// TIA Portal project "HydroPlantProject_V15.1" (V15.1) (continued)

   //EStop Alarm
   IF NOT "EStop" AND NOT "EStopAlarm" THEN
       "EStopAlarm" := 1;
       "EStopNotify" := 1;
   END_IF;

   IF "EStopAlarm" AND "AlarmReset" THEN
       "EStopAlarm" := 0;
       "EStopNotify" := 0;
   END_IF;

   IF "EStopNotify" AND "AlarmSilence" THEN
       "EStopNotify" := 0;
   END_IF;



   //Alarm Horn Control
   IF "FaultMode" AND NOT "AlarmHorn_Ctrl" THEN
       "AlarmHorn_Ctrl" := 1;
   END_IF;

   IF "AlarmHorn_Ctrl" AND ("AlarmReset" OR "AlarmSilence") THEN
       "AlarmHorn_Ctrl" := 0;
   END_IF;
END_FUNCTION_BLOCK

FUNCTION_BLOCK "ALARMS_STL"   // FB13, STL
{ S7_Optimized_Access := 'TRUE' }
VERSION : 0.1
   VAR
      OS1 : Bool;
      OS2 : Bool;
      OS3 : Bool;
      OS4 : Bool;
      OS5 : Bool;
      OS6 : Bool;
      OS7 : Bool;
      OS8 : Bool;
      OS9 : Bool;
      OS10 : Bool;
      OS11 : Bool;
      OS12 : Bool;
      OS13 : Bool;
      OS14 : Bool;
      OS15 : Bool;
      OS16 : Bool;
      OS17 : Bool;
   END_VAR
   VAR_TEMP
      ti1 : Time;
      ti2 : Time;
      ti3 : Time;
      ti4 : Time;
      ti5 : Time;
      ti6 : Time;
      ti7 : Time;
      t1 : Time;
      t2 : Time;
      t3 : Time;
      t4 : Time;
      t5 : Time;
      t6 : Time;
      t7 : Time;
      OILAT : Bool;
      OLFAT : Bool;
      OCAT : Bool;
      HOTAT : Bool;
      OSAT : Bool;
      HOFAT : Bool;
      BFAT : Bool;
   END_VAR
BEGIN

REGION Network 1
   //Oil Low Flow Alarm
         L     "OilFlow";
         L     "OilLLflowSp";
         <I;
         A     "OilPumpVFDen_Out";
         AN    "Brake_Out";
         JC    OLFtimer;
         CLR;
         A     "AlarmReset";
         FP    #OS1;
         JC    ResetOLFalarm;
         CLR;
         A     "AlarmSilence";
         FP    #OS2;
         JC    ResetOLFnotify;
         JU    OvercurrentAlarm;

   OLFtimer:CALL  "CONVERTTIME"
         ( Int1  := "OilLowFlowDelay_Sp",
           Time1 := #ti1
         );
         CALL  TON, "IEC_Timer_0_DB_18"
         ( IN := TRUE,
           PT := #ti1,
           Q  := #OLFAT,
           ET := #t1
         );
         A     #OLFAT;
         JC    SetOLFalarm;
         JU    OvercurrentAlarm;

   SetOLFalarm:SET;
         S     "OilLowFlowAlarm";
         S     "OilLowFlowNotify";
         JU    OvercurrentAlarm;

   ResetOLFalarm:R     "OilLowFlowAlarm";
         R     "OilLowFlowNotify";
         JU    OvercurrentAlarm;

   ResetOLFnotify:R     "OilLowFlowNotify";
         JU    OvercurrentAlarm;


   //Overcurrent Alarm
   OvercurrentAlarm:L     "Current";
         L     "OvercurrentSp";
         >I;
         JC    OCtimer;
         CLR;
         A     "AlarmReset";
         FP    #OS3;
         JC    ResetOCalarm;
         CLR;
         A     "AlarmSilence";
         FP    #OS4;
         JC    ResetOCnotify;
         JU    HighOilTempAlarm;

   OCtimer:CALL  "CONVERTTIME"
         ( Int1  := "OvercurrentDelay_Sp",
           Time1 := #ti2
         );
         CALL  TON, "IEC_Timer_0_DB_19"
         ( IN := true,
           PT := #ti2,
           Q  := #OCAT,
           ET := #t2
         );
         A     #OCAT;
         JC    SetOCalarm;
         JU    HighOilTempAlarm;

   SetOCalarm:SET;
         S     "OvercurrentAlarm";
         S     "OvercurrentNotify";
         JU    HighOilTempAlarm;

   ResetOCalarm:R     "OvercurrentAlarm";
         R     "OvercurrentNotify";
         JU    HighOilTempAlarm;

   ResetOCnotify:R     "OvercurrentNotify";
         JU    HighOilTempAlarm;


   //High Oil Temp Alarm
   HighOilTempAlarm:L     "OilTemp";
         L     "HighOilTempSp";
         >I;
         JC    HOTtimer;
         CLR;
         A     "AlarmReset";
         FP    #OS5;
         JC    ResetHOTalarm;
         CLR;
         A     "AlarmSilence";
         FP    #OS6;
         JC    ResetHOTnotify;
         JU    OverspeedAlarm;

   HOTtimer:CALL  "CONVERTTIME"
         ( Int1  := "HighOilTempDelay_Sp",
           Time1 := #ti3
         );
         CALL  TON, "IEC_Timer_0_DB_20"
         ( IN := TRUE,
           PT := #ti3,
           Q  := #HOTAT,
           ET := #t3
         );
         A     #HOTAT;
         JC    SetHOTalarm;
         JU    OverspeedAlarm;

   SetHOTalarm:SET;
         S     "HighOilTempAlarm";
         S     "HighOilTempNotify";
         JU    OverspeedAlarm;

   ResetHOTalarm:R     "HighOilTempAlarm";
         R     "HighOilTempNotify";
         JU    OverspeedAlarm;

   ResetHOTnotify:R     "HighOilTempNotify";
         JU    OverspeedAlarm;


   //Overspeed Alarm
   OverspeedAlarm:L     "RPM";
         L     "OverspeedSp";
         >I;
         JC    OStimer;
         CLR;
         A     "AlarmReset";
         FP    #OS7;
         JC    ResetOSalarm;
         CLR;
         A     "AlarmSilence";
         FP    #OS8;
         JC    ResetOSnotify;
         JU    HighOilFlowAlarm;

   OStimer:CALL  "CONVERTTIME"
         ( Int1  := "OverspeedDelay_Sp",
           Time1 := #ti4
         );
         CALL  TON, "IEC_Timer_0_DB_21"
         ( IN := TRUE,
           PT := #ti4,
           Q  := #OSAT,
           ET := #t4
         );
         A     #OSAT;
         JC    SetOSalarm;
         JU    HighOilFlowAlarm;

   SetOSalarm:SET;
         S     "OverspeedAlarm";
         S     "OverspeedNotify";
         JU    HighOilFlowAlarm;

   ResetOSalarm:R     "OverspeedAlarm";
         R     "OverspeedNotify";
         JU    HighOilFlowAlarm;

   ResetOSnotify:R     "OverspeedNotify";
         JU    HighOilFlowAlarm;


   //High Oil Flow Alarm
   HighOilFlowAlarm:L     "OilFlow";
         L     "OilHHflowSp";
         >I;
         JC    HOFtimer;
         CLR;
         A     "AlarmReset";
         FP    #OS9;
         JC    ResetHOFalarm;
         CLR;
         A     "AlarmSilence";
         FP    #OS10;
         JC    ResetHOFnotify;
         JU    BrakeFailureAlarm;

   HOFtimer:CALL  "CONVERTTIME"
         ( Int1  := "OilHighFlowDelay_Sp",
           Time1 := #ti5
         );
         CALL  TON, "IEC_Timer_0_DB_22"
         ( IN := TRUE,
           PT := #ti5,
           Q  := #HOFAT,
           ET := #t5
         );
         A     #HOFAT;
         JC    SetHOFalarm;
         JU    BrakeFailureAlarm;

   SetHOFalarm:SET;
         S     "OilHighFlowAlarm";
         S     "OilHighFlowNotify";
         JU    BrakeFailureAlarm;

   ResetHOFalarm:R     "OilHighFlowAlarm";
         R     "OilHighFlowNotify";
         JU    BrakeFailureAlarm;

   ResetHOFnotify:R     "OilHighFlowNotify";
         JU    BrakeFailureAlarm;


   //Brake Failure Alarm
   BrakeFailureAlarm:L     "RPM";
         L     0;
         >I;
         A     "Brake_Out";
         JC    BFtimer;
         CLR;
         A     "AlarmReset";
         FP    #OS11;
         JC    ResetBFalarm;
         CLR;
         A     "AlarmSilence";
         FP    #OS12;
         JC    ResetBFnotify;
         JU    EStoplarm;

   BFtimer:CALL  "CONVERTTIME"
         ( Int1  := "BrakeFailureDelay_Sp",
           Time1 := #ti6
         );
         CALL  TON, "IEC_Timer_0_DB_23"
         ( IN := TRUE,
           PT := #ti6,
           Q  := #BFAT,
           ET :=
         );
         A     #BFAT;
         JC    SetBFalarm;
         JU    EStoplarm;

   SetBFalarm:SET;
         S     "BrakeFailureAlarm";
         S     "BrakeFailureNotify";
         JU    EStoplarm;

   ResetBFalarm:R     "BrakeFailureAlarm";
         R     "BrakeFailureNotify";
         JU    EStoplarm;

   ResetBFnotify:R     "BrakeFailureNotify";
         JU    EStoplarm;


   //EStop Alarm
   EStoplarm:AN    "EStop";
         FP    #OS13;
         JC    SetESalarm;
         CLR;
         A     "AlarmReset";
         FP    #OS14;
         JC    ResetESalarm;
         CLR;
         A     "AlarmSilence";
         FP    #OS15;
         JC    ResetESnotify;
         JU    AlarmHornCtrl;

   SetESalarm:SET;
         S     "EStopAlarm";
         S     "EStopNotify";
         JU    AlarmHornCtrl;

   ResetESalarm:R     "EStopAlarm";
         R     "EStopNotify";
         JU    AlarmHornCtrl;

   ResetESnotify:R     "EStopNotify";
         JU    AlarmHornCtrl;



   //Alarm Horn Control
   AlarmHornCtrl:A     "FaultMode";
         FP    #OS16;
         JC    SetAlarmHorn;
         CLR;
         A     "AlarmReset";
         O     "AlarmSilence";
         FP    #OS17;
         JC    ResetAlarmHorn;
         JU    EndOfLine;

   SetAlarmHorn:SET;
         S     "AlarmHorn_Ctrl";
         JU    EndOfLine;

   ResetAlarmHorn:R     "AlarmHorn_Ctrl";
         JU    EndOfLine;



   EndOfLine:BE;
END_REGION
END_FUNCTION_BLOCK

FUNCTION_BLOCK "MODES_LAD"   // FB14, LAD
{ S7_Optimized_Access := 'TRUE' }
VERSION : 0.1
   VAR
      OS1 : Bool;
      OS2 : Bool;
      OS3 : Bool;
      OS4 : Bool;
      OS5 : Bool;
   END_VAR
   VAR_TEMP
      tv1 : Int;
      ti1 : Time;
      tv2 : Int;
      tv3 : Int;
      tv4 : Int;
      ti2 : Time;
      tv5 : Int;
      ti3 : Time;
   END_VAR
   VAR_TEMP   // added for the SCL form of the ladder/FBD networks
      _w1 : Bool;
      _w2 : Bool;
      _w3 : Bool;
   END_VAR
BEGIN

REGION Network 1
   // Warmup Mode
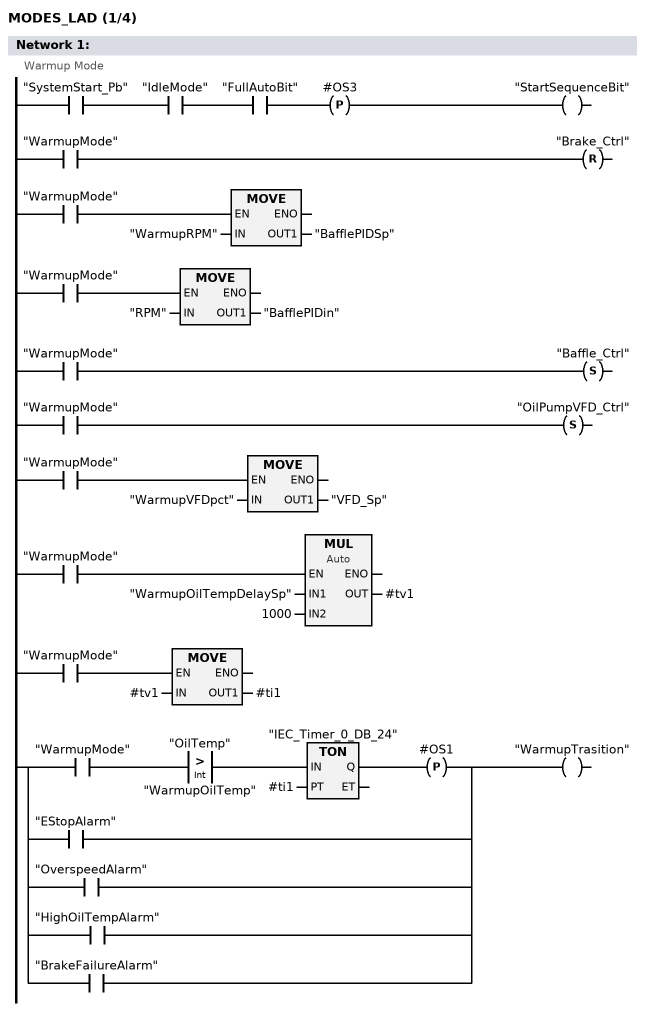
   #_w1 := "SystemStart_Pb" AND "IdleMode" AND "FullAutoBit";
   #_w2 := #_w1 AND NOT #OS3;   // rising edge
   #OS3 := #_w1;
   "StartSequenceBit" := #_w2;
   IF "WarmupMode" THEN
       "Brake_Ctrl" := FALSE;
       "BafflePIDSp" := "WarmupRPM";
       "BafflePIDin" := "RPM";
       "Baffle_Ctrl" := TRUE;
       "OilPumpVFD_Ctrl" := TRUE;
       "VFD_Sp" := "WarmupVFDpct";
       #tv1 := "WarmupOilTempDelaySp" * 1000;
       #ti1 := #tv1;
   END_IF;
   "IEC_Timer_0_DB_24".TON(IN := "WarmupMode" AND ("OilTemp" > "WarmupOilTemp"), PT := #ti1);
   #_w3 := "IEC_Timer_0_DB_24".Q AND NOT #OS1;   // rising edge
   #OS1 := "IEC_Timer_0_DB_24".Q;
   "WarmupTrasition" := #_w3 OR "EStopAlarm" OR "OverspeedAlarm" OR "HighOilTempAlarm" OR "BrakeFailureAlarm";
END_REGION

REGION Network 2
   // Stabilize Mode
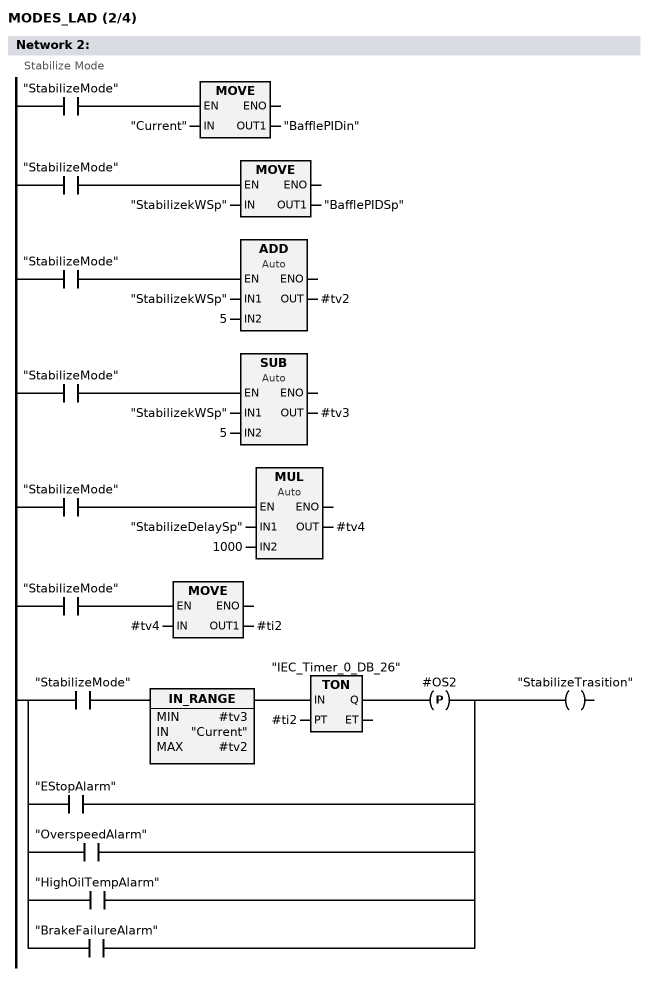
   IF "StabilizeMode" THEN
       "BafflePIDin" := "Current";
       "BafflePIDSp" := "StabilizekWSp";
       #tv2 := "StabilizekWSp" + 5;
       #tv3 := "StabilizekWSp" - 5;
       #tv4 := "StabilizeDelaySp" * 1000;
       #ti2 := #tv4;
   END_IF;
   "IEC_Timer_0_DB_26".TON(IN := "StabilizeMode" AND (#tv3 <= "Current") AND ("Current" <= #tv2), PT := #ti2);
   #_w1 := "IEC_Timer_0_DB_26".Q AND NOT #OS2;   // rising edge
   #OS2 := "IEC_Timer_0_DB_26".Q;
   "StabilizeTrasition" := #_w1 OR "EStopAlarm" OR "OverspeedAlarm" OR "HighOilTempAlarm" OR "BrakeFailureAlarm";
END_REGION

REGION Network 3
   // Generation Mode
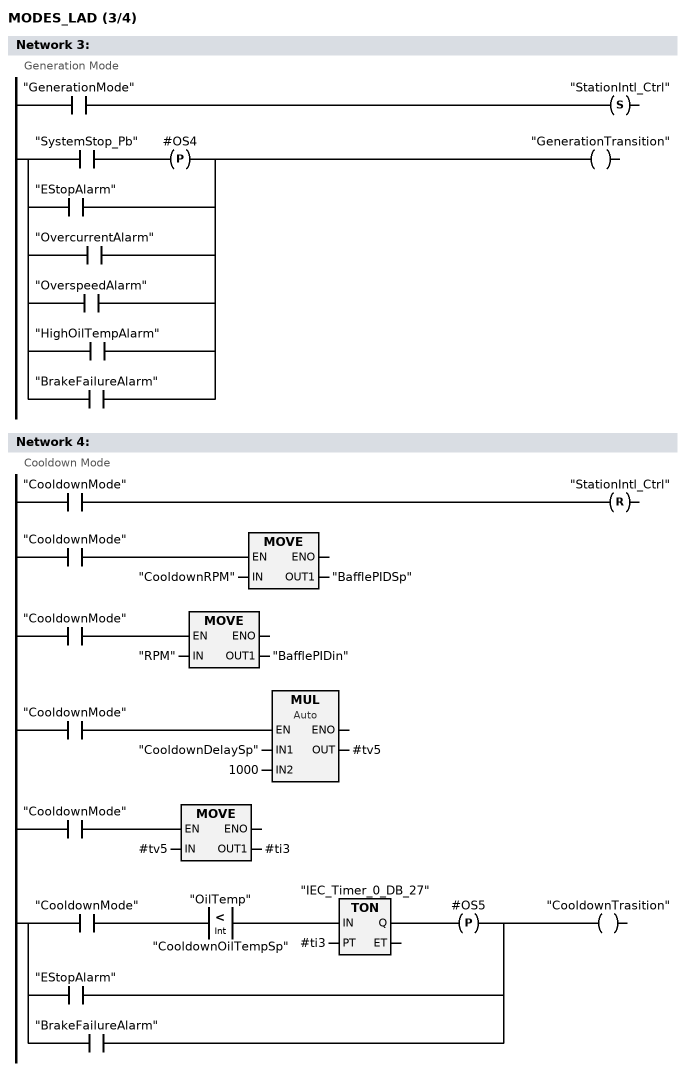
   RUNG wire#powerrail
      Contact( "GenerationMode" )
      S_Coil( "StationIntl_Ctrl" )
   END_RUNG
   RUNG wire#powerrail
      Contact( "SystemStop_Pb" )
      P_Trig( #OS4 )
      wire#w1
      Coil( "GenerationTransition" )
   END_RUNG
   RUNG wire#powerrail
      Contact( "EStopAlarm" )
   END_RUNG wire#w1
   RUNG wire#powerrail
      Contact( "OvercurrentAlarm" )
   END_RUNG wire#w1
   RUNG wire#powerrail
      Contact( "OverspeedAlarm" )
   END_RUNG wire#w1
   RUNG wire#powerrail
      Contact( "HighOilTempAlarm" )
   END_RUNG wire#w1
   RUNG wire#powerrail
      Contact( "BrakeFailureAlarm" )
   END_RUNG wire#w1
   // the same network as SCL:
   IF "GenerationMode" THEN "StationIntl_Ctrl" := TRUE; END_IF;
   #_w1 := "SystemStop_Pb" AND NOT #OS4;   // rising edge
   #OS4 := "SystemStop_Pb";
   "GenerationTransition" := #_w1 OR "EStopAlarm" OR "OvercurrentAlarm" OR "OverspeedAlarm" OR "HighOilTempAlarm" OR "BrakeFailureAlarm";
END_REGION

REGION Network 4
   // Cooldown Mode
   IF "CooldownMode" THEN
       "StationIntl_Ctrl" := FALSE;
       "BafflePIDSp" := "CooldownRPM";
       "BafflePIDin" := "RPM";
       #tv5 := "CooldownDelaySp" * 1000;
       #ti3 := #tv5;
   END_IF;
   "IEC_Timer_0_DB_27".TON(IN := "CooldownMode" AND ("OilTemp" < "CooldownOilTempSp"), PT := #ti3);
   #_w1 := "IEC_Timer_0_DB_27".Q AND NOT #OS5;   // rising edge
   #OS5 := "IEC_Timer_0_DB_27".Q;
   "CooldownTrasition" := #_w1 OR "EStopAlarm" OR "BrakeFailureAlarm";
END_REGION

REGION Network 5
   // Idle Mode
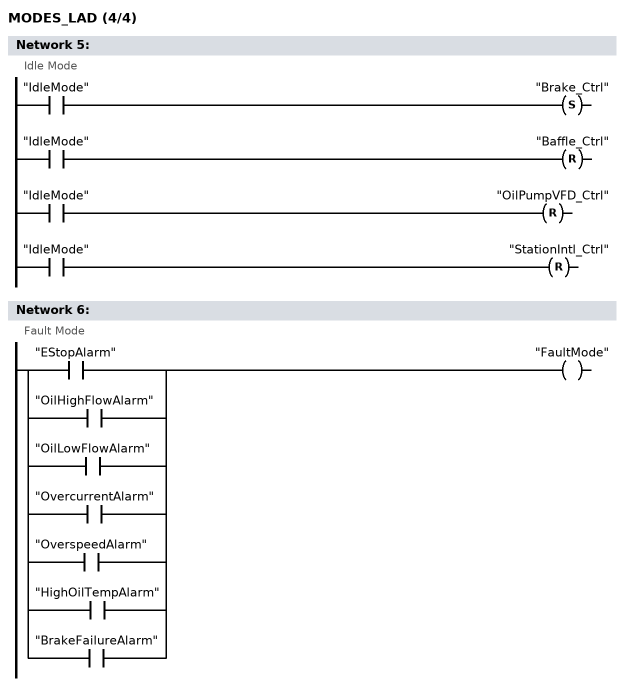
   RUNG wire#powerrail
      Contact( "IdleMode" )
      S_Coil( "Brake_Ctrl" )
   END_RUNG
   RUNG wire#powerrail
      Contact( "IdleMode" )
      R_Coil( "Baffle_Ctrl" )
   END_RUNG
   RUNG wire#powerrail
      Contact( "IdleMode" )
      R_Coil( "OilPumpVFD_Ctrl" )
   END_RUNG
   RUNG wire#powerrail
      Contact( "IdleMode" )
      R_Coil( "StationIntl_Ctrl" )
   END_RUNG
   // the same network as SCL:
   IF "IdleMode" THEN
       "Brake_Ctrl" := TRUE;
       "Baffle_Ctrl" := FALSE;
       "OilPumpVFD_Ctrl" := FALSE;
       "StationIntl_Ctrl" := FALSE;
   END_IF;
END_REGION

REGION Network 6
   // Fault Mode
   RUNG wire#powerrail
      Contact( "EStopAlarm" )
      wire#w1
      Coil( "FaultMode" )
   END_RUNG
   RUNG wire#powerrail
      Contact( "OilHighFlowAlarm" )
   END_RUNG wire#w1
   RUNG wire#powerrail
      Contact( "OilLowFlowAlarm" )
   END_RUNG wire#w1
   RUNG wire#powerrail
      Contact( "OvercurrentAlarm" )
   END_RUNG wire#w1
   RUNG wire#powerrail
      Contact( "OverspeedAlarm" )
   END_RUNG wire#w1
   RUNG wire#powerrail
      Contact( "HighOilTempAlarm" )
   END_RUNG wire#w1
   RUNG wire#powerrail
      Contact( "BrakeFailureAlarm" )
   END_RUNG wire#w1
   // the same network as SCL:
   "FaultMode" := "EStopAlarm" OR "OilHighFlowAlarm" OR "OilLowFlowAlarm" OR "OvercurrentAlarm" OR "OverspeedAlarm" OR "HighOilTempAlarm" OR "BrakeFailureAlarm";
END_REGION
END_FUNCTION_BLOCK

FUNCTION_BLOCK "MODES_FBD"   // FB15, FBD
{ S7_Optimized_Access := 'TRUE' }
VERSION : 0.1
   VAR
      OS1 : Bool;
      OS2 : Bool;
      OS3 : Bool;
      OS4 : Bool;
      OS5 : Bool;
   END_VAR
   VAR_TEMP
      ti1 : Time;
      tv1 : Int;
      tv2 : Int;
      ti3 : Time;
      ti2 : Time;
   END_VAR
   VAR_TEMP   // added for the SCL form of the ladder/FBD networks
      _w1 : Bool;
      _w2 : Bool;
      _w3 : Bool;
   END_VAR
BEGIN

REGION Network 1
   // Warmup Mode
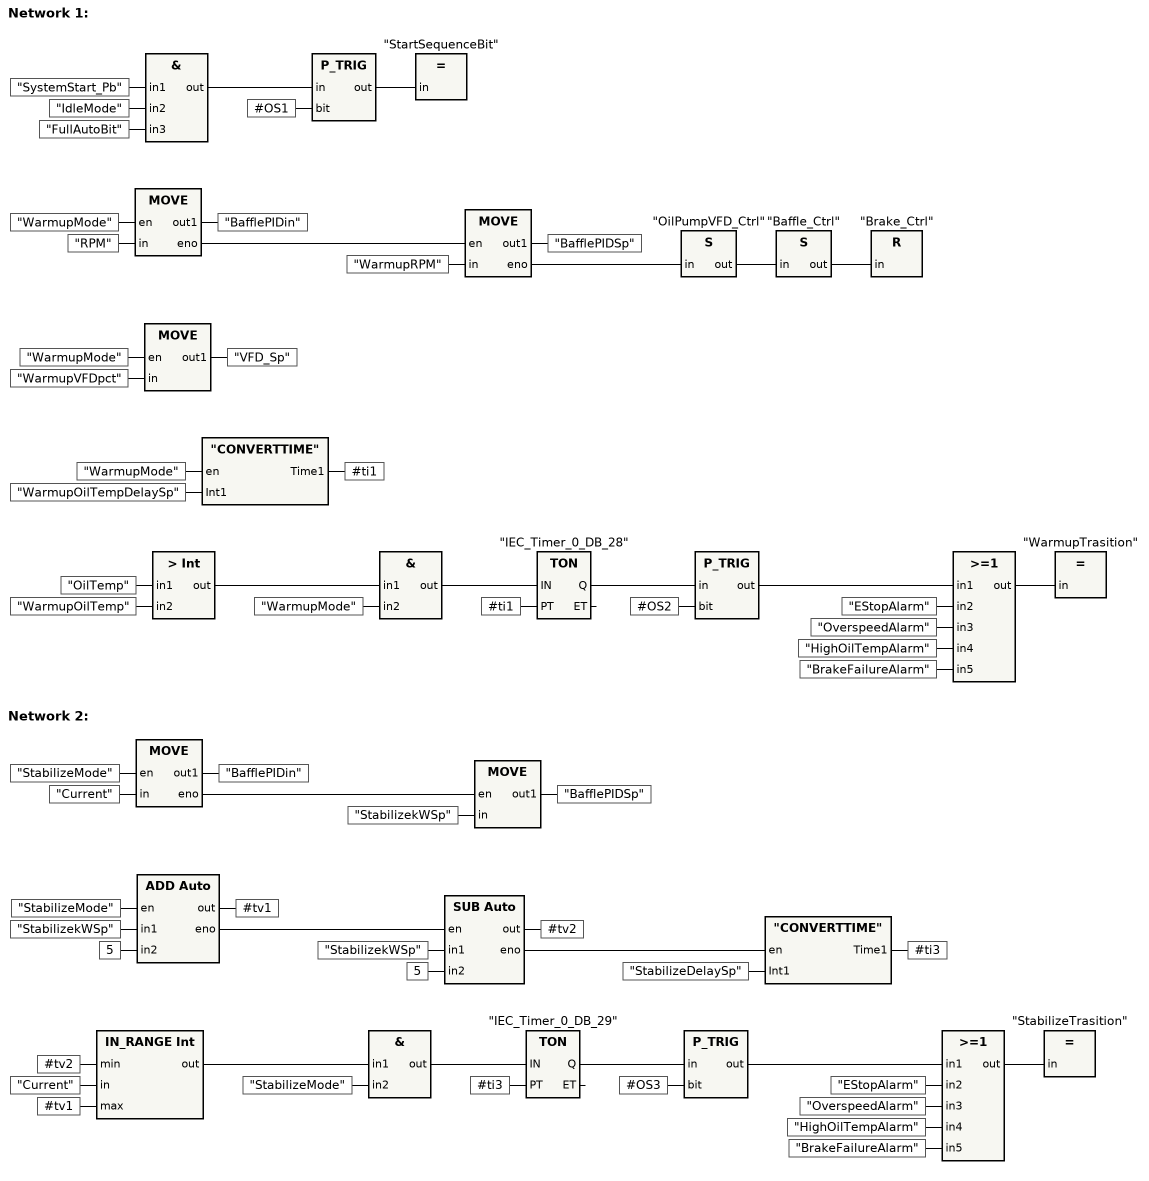
   #_w1 := "SystemStart_Pb" AND "IdleMode" AND "FullAutoBit";
   #_w2 := #_w1 AND NOT #OS1;   // rising edge
   #OS1 := #_w1;
   "StartSequenceBit" := #_w2;
   IF "WarmupMode" THEN
       "BafflePIDin" := "RPM";
       "BafflePIDSp" := "WarmupRPM";
       "OilPumpVFD_Ctrl" := TRUE;
       "Baffle_Ctrl" := TRUE;
       "Brake_Ctrl" := FALSE;
       "VFD_Sp" := "WarmupVFDpct";
       "CONVERTTIME"(Int1 := "WarmupOilTempDelaySp", Time1 => #ti1);
   END_IF;
   "IEC_Timer_0_DB_28".TON(IN := ("OilTemp" > "WarmupOilTemp") AND "WarmupMode", PT := #ti1);
   #_w3 := "IEC_Timer_0_DB_28".Q AND NOT #OS2;   // rising edge
   #OS2 := "IEC_Timer_0_DB_28".Q;
   "WarmupTrasition" := #_w3 OR "EStopAlarm" OR "OverspeedAlarm" OR "HighOilTempAlarm" OR "BrakeFailureAlarm";
END_REGION

REGION Network 2
   // Stabilize Mode
   IF "StabilizeMode" THEN
       "BafflePIDin" := "Current";
       "BafflePIDSp" := "StabilizekWSp";
       #tv1 := "StabilizekWSp" + 5;
       #tv2 := "StabilizekWSp" - 5;
       "CONVERTTIME"(Int1 := "StabilizeDelaySp", Time1 => #ti3);
   END_IF;
   "IEC_Timer_0_DB_29".TON(IN := (#tv2 <= "Current") AND ("Current" <= #tv1) AND "StabilizeMode", PT := #ti3);
   #_w1 := "IEC_Timer_0_DB_29".Q AND NOT #OS3;   // rising edge
   #OS3 := "IEC_Timer_0_DB_29".Q;
   "StabilizeTrasition" := #_w1 OR "EStopAlarm" OR "OverspeedAlarm" OR "HighOilTempAlarm" OR "BrakeFailureAlarm";
END_REGION

REGION Network 3
   // Generation Mode
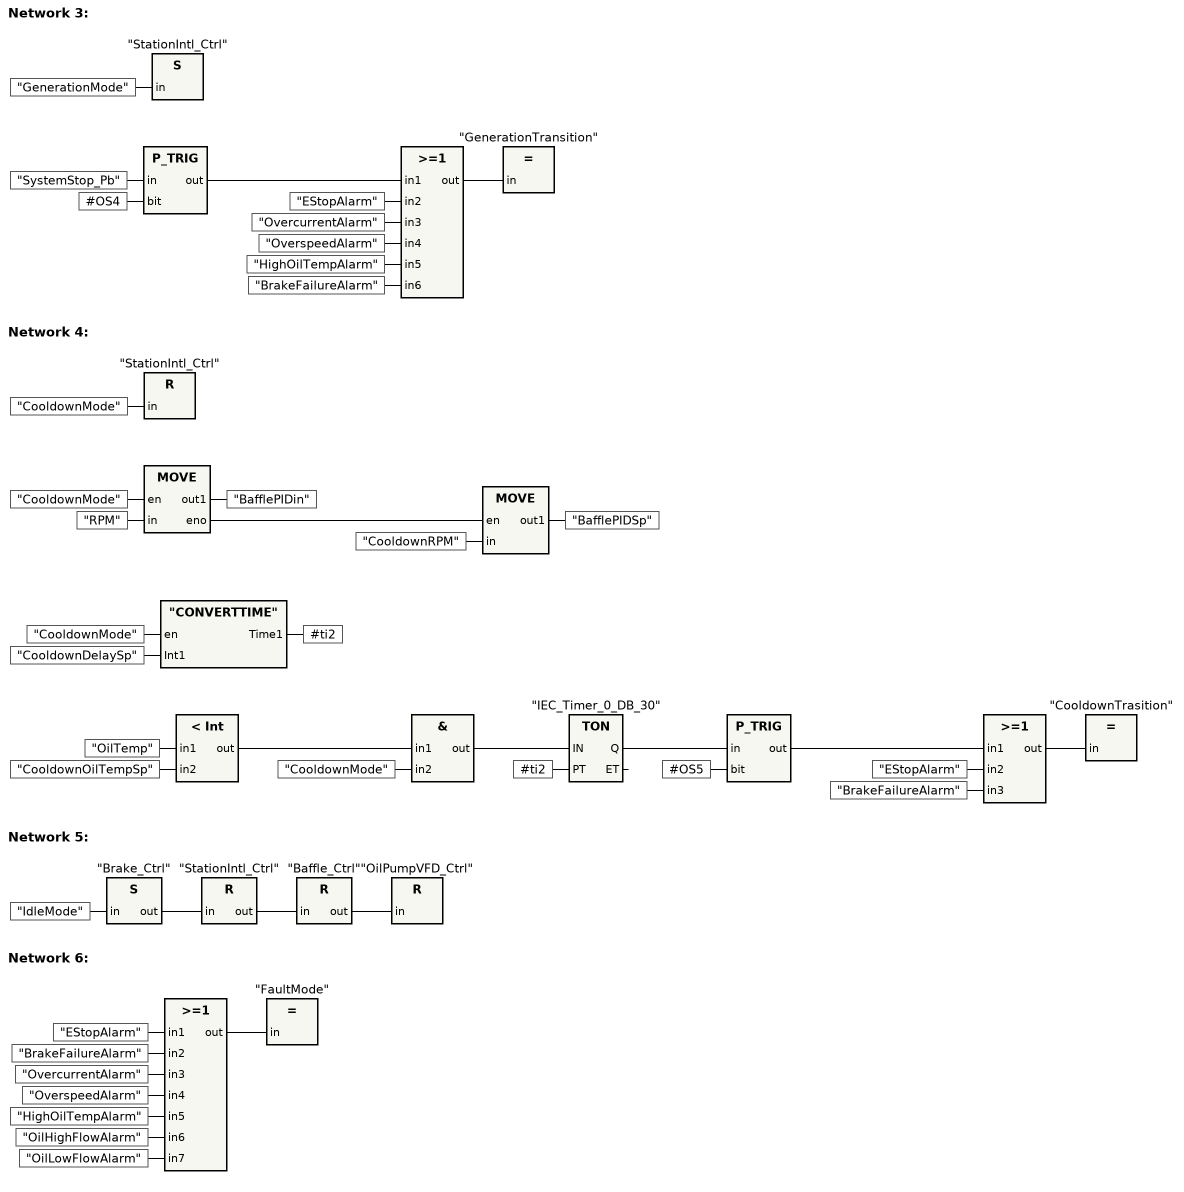
   IF "GenerationMode" THEN "StationIntl_Ctrl" := TRUE; END_IF;
   #_w1 := "SystemStop_Pb" AND NOT #OS4;   // rising edge
   #OS4 := "SystemStop_Pb";
   "GenerationTransition" := #_w1 OR "EStopAlarm" OR "OvercurrentAlarm" OR "OverspeedAlarm" OR "HighOilTempAlarm" OR "BrakeFailureAlarm";
END_REGION

REGION Network 4
   // Cooldown Mode
   IF "CooldownMode" THEN
       "StationIntl_Ctrl" := FALSE;
       "BafflePIDin" := "RPM";
       "BafflePIDSp" := "CooldownRPM";
       "CONVERTTIME"(Int1 := "CooldownDelaySp", Time1 => #ti2);
   END_IF;
   "IEC_Timer_0_DB_30".TON(IN := ("OilTemp" < "CooldownOilTempSp") AND "CooldownMode", PT := #ti2);
   #_w1 := "IEC_Timer_0_DB_30".Q AND NOT #OS5;   // rising edge
   #OS5 := "IEC_Timer_0_DB_30".Q;
   "CooldownTrasition" := #_w1 OR "EStopAlarm" OR "BrakeFailureAlarm";
END_REGION

REGION Network 5
   // Idle Mode
   IF "IdleMode" THEN
       "Brake_Ctrl" := TRUE;
       "StationIntl_Ctrl" := FALSE;
       "Baffle_Ctrl" := FALSE;
       "OilPumpVFD_Ctrl" := FALSE;
   END_IF;
END_REGION

REGION Network 6
   // Fault Mode
   "FaultMode" := "EStopAlarm" OR "BrakeFailureAlarm" OR "OvercurrentAlarm" OR "OverspeedAlarm" OR "HighOilTempAlarm" OR "OilHighFlowAlarm" OR "OilLowFlowAlarm";
END_REGION
END_FUNCTION_BLOCK

FUNCTION_BLOCK "MODES_SCL"   // FB16, SCL
{ S7_Optimized_Access := 'TRUE' }
VERSION : 0.1
   VAR_TEMP
      ti1 : Time;
      ti2 : Time;
      tv1 : Int;
      tv2 : Int;
      ti3 : Time;
      warmupdelaytrigger : Bool;
      stabilizedelaytrigger : Bool;
      ti4 : Time;
      ti5 : Time;
      cooldowndelaytrigger : Bool;
      ti6 : Time;
   END_VAR
BEGIN
   //EStop Handling
   IF "EStopAlarm" OR "BrakeFailureAlarm" THEN
       "WarmupTrasition" := 1;
       "StabilizeTrasition" := 1;
       "GenerationTransition" := 1;
       "CooldownTrasition" := 1;
   ELSE
       "WarmupTrasition" := 0;
       "StabilizeTrasition" := 0;
       "GenerationTransition" := 0;
       "CooldownTrasition" := 0;

       //Warmup Mode
       IF "SystemStart_Pb" AND "IdleMode" AND "FullAutoBit" THEN
           "StartSequenceBit" := 1;
       ELSE
           "StartSequenceBit" := 0;
       END_IF;


       IF "WarmupMode" THEN
           "Brake_Ctrl" := 0;
           "BafflePIDin" := "RPM";
           "BafflePIDSp" := "WarmupRPM";
           "VFD_Sp" := "WarmupVFDpct";
           IF "OilTemp" > "WarmupOilTemp" THEN
               "CONVERTTIME"(Int1 := "WarmupOilTempDelaySp",
                             Time1 => #ti1);
               "IEC_Timer_0_DB_31".TON(IN := TRUE,
                                       PT := #ti1,
                                       Q => #warmupdelaytrigger,
                                       ET => #ti2);
           ELSE
               RESET_TIMER("IEC_Timer_0_DB_31");
           END_IF;
           IF #warmupdelaytrigger THEN
               RESET_TIMER("IEC_Timer_0_DB_31");
               "WarmupTrasition" := 1;
           END_IF;
       ELSE
           "WarmupTrasition" := 0;
       END_IF;

       IF "OverspeedAlarm" OR "HighOilTempAlarm" THEN
           "WarmupTrasition" := 1;
       END_IF;

       //Stabilize Mode
       IF "StabilizeMode" THEN
           "BafflePIDin" := "Current";
           "BafflePIDSp" := "StabilizekWSp";
           #tv1 := "StabilizekWSp" - 5;
           #tv2 := "StabilizekWSp" + 5;
           IF "Current" < #tv2 AND "Current" > #tv1 THEN
               "CONVERTTIME"(Int1 := "StabilizeDelaySp",
                             Time1 => #ti3);
               "IEC_Timer_0_DB_32".TON(IN := TRUE,
                                       PT := #ti3,
                                       Q => #stabilizedelaytrigger,
                                       ET => #ti4);
           ELSE
               RESET_TIMER("IEC_Timer_0_DB_32");
           END_IF;
           IF #stabilizedelaytrigger THEN
               RESET_TIMER("IEC_Timer_0_DB_31");
               "StabilizeTrasition" := 1;
           END_IF;
       ELSE
           "StabilizeTrasition" := 0;
       END_IF;

       IF "OverspeedAlarm" OR "HighOilTempAlarm" THEN
           "StabilizeTrasition" := 1;
       END_IF;


       //Generation Mode
       IF "GenerationMode" THEN
           "StationIntl_Ctrl" := 1;
           IF "SystemStop_Pb" THEN
               "GenerationTransition" := 1;
           END_IF;
       ELSE
           "GenerationTransition" := 0;
       END_IF;

       IF "OvercurrentAlarm" OR "OverspeedAlarm" OR "HighOilTempAlarm" THEN
           "GenerationTransition" := 1;
       END_IF;


       //Cooldown Mode
       IF "CooldownMode" THEN
           "StationIntl_Ctrl" := 0;
           "BafflePIDin" := "RPM";
           "BafflePIDSp" := "CooldownRPMSp";
           IF "OilTemp" < "CooldownOilTempSp" THEN
               "CONVERTTIME"(Int1 := "CooldownDelaySp",
                             Time1 => #ti5);
               "IEC_Timer_0_DB_33".TON(IN := TRUE,
                                       PT := #ti5,
                                       Q => #cooldowndelaytrigger,
                                       ET => #ti6);
           ELSE
               RESET_TIMER("IEC_Timer_0_DB_33");
           END_IF;
           IF #cooldowndelaytrigger THEN
               RESET_TIMER("IEC_Timer_0_DB_33");
               "CooldownTrasition" := 1;
           END_IF;
       ELSE
           "CooldownTrasition" := 0;
       END_IF;


       //Fault Mode
       IF "EStopAlarm" OR "BrakeFailureAlarm" OR "OvercurrentAlarm" OR "OverspeedAlarm" OR "HighOilTempAlarm" OR "OilHighFlowAlarm" OR "OilLowFlowAlarm" THEN
           "FaultMode" := 1;
       ELSE
           "FaultMode" := 0;
       END_IF;

   END_IF;

   //Idle Mode
   IF "IdleMode" THEN
       "Brake_Ctrl" := 1;
       "OilPumpVFD_Ctrl" := 0;
       "Baffle_Ctrl" := 0;
       "StationIntl_Ctrl" := 0;
   END_IF;
END_FUNCTION_BLOCK

FUNCTION_BLOCK "MODES_STL"   // FB17, STL
{ S7_Optimized_Access := 'TRUE' }
VERSION : 0.1
   VAR
      OS1 : Bool;
      OS2 : Bool;
   END_VAR
   VAR_TEMP
      ti1 : Time;
      warmupdelaytrigger : Bool;
      ti2 : Time;
      tv1 : Int;
      tv2 : Int;
      tb1 : Bool;
      ti3 : Time;
      stabilizedelaytrigger : Bool;
      ti4 : Time;
      ti5 : Time;
      ti6 : Time;
      cooldowndelaytrigger : Bool;
   END_VAR
BEGIN

REGION Network 1
   //EStop Handling
   EStop:A     "EStopAlarm";
         O     "BrakeFailureAlarm";
         JC    EStopTransitions;
         JU    ResetTransitions;

   EStopTransitions:SET;
         S     "WarmupTrasition";
         S     "StabilizeTrasition";
         S     "GenerationTransition";
         S     "CooldownTrasition";
         JU    JumpToMode;

   ResetTransitions:CLR;
         NOT;
         R     "WarmupTrasition";
         R     "StabilizeTrasition";
         R     "GenerationTransition";
         R     "CooldownTrasition";
         JU    JumpToMode;

   JumpToMode:A     "WarmupMode";
         JC    StartWarmup;
         CLR;
         A     "StabilizeMode";
         JC    StabilizeMode;
         CLR;
         A     "GenerationMode";
         JC    GenerationMode;
         CLR;
         A     "CooldownMode";
         JC    CooldownMode;
         CLR;
         A     "IdleMode";
         JC    IdleMode;
         JU    EndOfLine;

   //Warmup Mode
   StartWarmup:SET;
         R     "WarmupTrasition";
         R     "StabilizeTrasition";
         R     "GenerationTransition";
         R     "CooldownTrasition";
         R     "StartSequenceBit";
         CLR;
         A     "WarmupMode";
         JC    WarmupMode;
         CLR;
         A     "StabilizeMode";
         JC    StabilizeMode;
         CLR;
         A     "GenerationMode";
         JC    GenerationMode;
         CLR;
         A     "CooldownMode";
         JC    CooldownMode;
         CLR;
         A     "IdleMode";
         JC    IdleMode;
         JU    EndOfLine;

   WarmupMode:SET;
         NOT;
         R     "Brake_Ctrl";
         L     "WarmupRPM";
         T     "BafflePIDSp";
         L     "RPM";
         T     "BafflePIDin";

         SET;
         S     "OilPumpVFD_Ctrl";
         S     "Baffle_Ctrl";
         L     "WarmupVFDpct";
         T     "VFD_Sp";

         L     "OilTemp";
         L     "WarmupOilTemp";
         >I;
         JC    WarmupTime;
         CALL  RESET_TIMER
         ( "TIMER" := "IEC_Timer_0_DB_34"
         );
         JU    StabilizeMode;

   WarmupTime:CALL  "CONVERTTIME"
         ( Int1  := "WarmupOilTempDelaySp",
           Time1 := #ti1
         );
         CALL  TON, "IEC_Timer_0_DB_34"
         ( IN := TRUE,
           PT := #ti1,
           Q  := #warmupdelaytrigger,
           ET := #ti2
         );
         A     #warmupdelaytrigger;
         JC    WarmupExit;
         CLR;
         A     "OverspeedAlarm";
         O     "HighOilTempAlarm";
         JC    WarmupExit;
         JU    StabilizeMode;

   WarmupExit:S     "WarmupTrasition";
         CALL  RESET_TIMER
         ( "TIMER" := "IEC_Timer_0_DB_34"
         );
         JU    StabilizeMode;

   //Stabilize Mode
   StabilizeMode:SET;
         NOT;
         R     "WarmupTrasition";
         L     "StabilizekWSp";
         T     "BafflePIDSp";
         L     "Current";
         T     "BafflePIDin";
         L     "StabilizekWSp";
         L     5;
         +I;
         T     #tv1;
         L     "StabilizekWSp";
         L     5;
         -I;
         T     #tv2;
         L     "Current";
         L     #tv1;
         <I;
         S     #tb1;
         L     "Current";
         L     #tv2;
         >I;
         A     #tb1;
         JC    StabilizeTime;
         CALL  RESET_TIMER
         ( "TIMER" := "IEC_Timer_0_DB_35"
         );
         JU    GenerationMode;

   StabilizeTime:CALL  "CONVERTTIME"
         ( Int1  := "StabilizeDelaySp",
           Time1 := #ti3
         );
         CALL  TON , "IEC_Timer_0_DB_35"
         ( IN := TRUE,
           PT := #ti3,
           Q  := #stabilizedelaytrigger,
           ET := #ti4
         );
         A     #stabilizedelaytrigger;
         JC    StabilizeExit;
         CLR;
         A     "OverspeedAlarm";
         O     "HighOilTempAlarm";
         JC    StabilizeExit;
         JU    GenerationMode;

   StabilizeExit:S     "StabilizeTrasition";
         CALL  RESET_TIMER
         ( "TIMER" := "IEC_Timer_0_DB_35"
         );
         JU    GenerationMode;

   //Generation Mode
   GenerationMode:SET;
         NOT;
         R     "StabilizeTrasition";
         SET;
         S     "StationIntl_Ctrl";
         A     "SystemStop_Pb";
         JC    GenerationExit;
         CLR;
         A     "OvercurrentAlarm";
         JC    GenerationExit;
         CLR;
         A     "OverspeedAlarm";
         O     "HighOilTempAlarm";
         JC    GenerationExit;
         JU    CooldownMode;

   GenerationExit:S     "GenerationTransition";
         JU    CooldownMode;

   // Cooldown Mode
   CooldownMode:SET;
         NOT;
         R     "GenerationTransition";
         R     "StationIntl_Ctrl";
         L     "CooldownRPM";
         T     "BafflePIDSp";
         L     "RPM";
         T     "BafflePIDin";
         L     "OilTemp";
         L     "CooldownOilTempSp";
         <I;
         JC    CooldownTime;
         CALL  RESET_TIMER
         ( "TIMER" := "IEC_Timer_0_DB_36"
         );
         JU    IdleMode;

   CooldownTime:CALL  "CONVERTTIME"
         ( Int1  := "CooldownDelaySp",
           Time1 := #ti5
         );
         CALL  TON , "IEC_Timer_0_DB_36"
         ( IN := TRUE,
           PT := #ti5,
           Q  := #cooldowndelaytrigger,
           ET := #ti6
         );
         A     #cooldowndelaytrigger;
         JC    CooldownExit;
         JU    IdleMode;

   CooldownExit:S     "CooldownTrasition";
         CALL  RESET_TIMER
         ( "TIMER" := "IEC_Timer_0_DB_36"
         );
         JU    IdleMode;


   //Idle Mode
   IdleMode:SET;
         NOT;
         R     "CooldownTrasition";
         R     "StationIntl_Ctrl";
         S     "Brake_Ctrl";
         R     "Baffle_Ctrl";
         R     "OilPumpVFD_Ctrl";
         CLR;
         A     "SystemStart_Pb";
         A     "IdleMode";
         A     "FullAutoBit";
         FP    #OS1;
         S     "StartSequenceBit";
         JU    EndOfLine;

   //Fault Mode
   EndOfLine:A     "EStopAlarm";
         O     "BrakeFailureAlarm";
         O     "OvercurrentAlarm";
         O     "OverspeedAlarm";
         O     "HighOilTempAlarm";
         O     "OilHighFlowAlarm";
         O     "OilLowFlowAlarm";
         =     "FaultMode";
END_REGION
END_FUNCTION_BLOCK

FUNCTION_BLOCK "SEQUENCE"   // FB18, GRAPH_PLUS
{ S7_Optimized_Access := 'TRUE' }
VERSION : 0.1
   VAR_INPUT
      OFF_SQ : Bool := false;   // Turn sequence off
      INIT_SQ : Bool := false;   // Set sequence to initial state
      ACK_EF : Bool := false;   // Acknowledge all errors and faults
      S_PREV : Bool := false;   // Output previous step in parameter S_NO
      S_NEXT : Bool := false;   // Indicate next step in parameter S_NO
      SW_AUTO : Bool := false;   // Automatic mode
      SW_TAP : Bool := false;   // Semiautomatic/switch with transition
      SW_TOP : Bool := false;   // Semiautomatic/ignore transition
      SW_MAN : Bool := false;   // Manual mode
      S_SEL : Int := 0;   // Select step to be output to S_NO
      S_ON : Bool := false;   // Activate step indicated in S_NO
      S_OFF : Bool := false;   // Deactivate step indicated S_NO
      T_PUSH : Bool := false;   // Enable transition to switch in semi automatic mode
   END_VAR
   VAR_OUTPUT
      S_NO : Int := 0;   // Step number
      S_MORE : Bool := false;   // More steps are available and can be shown in S_NO
      S_ACTIVE : Bool := false;   // Step indicated in S_NO is active
      ERR_FLT : Bool := false;   // Interlock or supervision group error
      AUTO_ON : Bool := false;   // Automatic mode is active
      TAP_ON : Bool := false;   // Semiautomatic mode/step with transition enabled
      TOP_ON : Bool := false;   // Semiautomatic mode/ignore transition enabled
      MAN_ON : Bool := false;   // Manual mode is active
   END_VAR
   VAR
      HMI_INFO : Array[0..8] of UInt;
      IF_PAR : G7_IfParPlus_V2;
      RT_DATA : G7_RTDataPlus_V2;   // Internal data area
      Trans1 : G7_TransitionPlus_V2;   // Transition structure
      Trans2 : G7_TransitionPlus_V2;   // Transition structure
      Trans3 : G7_TransitionPlus_V2;   // Transition structure
      Trans4 : G7_TransitionPlus_V2;   // Transition structure
      Trans5 : G7_TransitionPlus_V2;   // Transition structure
      Idle : G7_StepPlus_V2;   // Step structure
      Warmup : G7_StepPlus_V2;   // Step structure
      Stabilize : G7_StepPlus_V2;   // Step structure
      Generation : G7_StepPlus_V2;   // Step structure
      Cooldown : G7_StepPlus_V2;   // Step structure
      SINI : Array[0..1] of USInt;
      LSTT : Array[0..4] of USInt;
      ATAJ : Array[0..4] of USInt;
      ATAB : Array[0..4] of USInt;
      PSTT : Array[0..4] of USInt;
      NSTT : Array[0..4] of USInt;
      ASSJ : Array[0..4] of USInt;
      ASSB : Array[0..4] of USInt;
      PTTS : Array[0..4] of USInt;
      NTTS : Array[0..4] of USInt;
      SW_SQTS : Array[0..4] of USInt;
      SWITCH : Array[0..0] of USInt;
      TVX : Array[0..1] of USInt;
      TTX : Array[0..1] of USInt;
      TSX : Array[0..1] of USInt;
      S00X : Array[0..1] of USInt;
      SOFFX : Array[0..1] of USInt;
      SONX : Array[0..1] of USInt;
      SAX : Array[0..1] of USInt;
      SERRX : Array[0..5] of USInt;
      SMX : Array[0..5] of USInt;
      S0X : Array[0..5] of USInt;
      S1X : Array[0..5] of USInt;
      IL_ALARM_INST : Program_Alarm;
      SUP_ALARM_INST : Program_Alarm;
      STEP_TIME_ALARM_INST : Program_Alarm;
      IEC_TIMER_INST : IEC_TIMER;
      TRANSACTION_FLAG : Bool := false;
   END_VAR
   // SINI[0] := 2;
   // SINI[1] := 1;
   // LSTT[0] := 255;
   // LSTT[1] := 255;
   // LSTT[2] := 255;
   // LSTT[4] := 255;
   // ATAJ[1] := 1;
   // ATAJ[2] := 2;
   // ATAJ[3] := 3;
   // ATAJ[4] := 4;
   // ATAB[1] := 1;
   // ATAB[2] := 2;
   // ATAB[3] := 3;
   // ATAB[4] := 4;
   // PSTT[0] := 1;
   // PSTT[1] := 2;
   // PSTT[2] := 3;
   // PSTT[3] := 4;
   // NSTT[0] := 2;
   // NSTT[1] := 3;
   // NSTT[2] := 4;
   // NSTT[4] := 1;
   // ASSJ[1] := 1;
   // ASSJ[2] := 2;
   // ASSJ[3] := 3;
   // ASSJ[4] := 4;
   // ASSB[1] := 1;
   // ASSB[2] := 2;
   // ASSB[3] := 3;
   // ASSB[4] := 4;
   // PTTS[0] := 255;
   // PTTS[1] := 4;
   // PTTS[3] := 1;
   // PTTS[4] := 2;
   // NTTS[0] := 4;
   // NTTS[2] := 1;
   // NTTS[3] := 2;
   // NTTS[4] := 3;
   // TVX[0] := 16#1;
   // TTX[0] := 16#1;
   // TSX[0] := 16#1;
   // S00X[0] := 16#1;
   // SOFFX[0] := 16#1;
   // SONX[0] := 16#1;
   // SAX[0] := 16#1;
   // SERRX[0] := 16#1;
   // SMX[0] := 16#1;
   // S0X[0] := 16#1;
   // S1X[0] := 16#1;
BEGIN
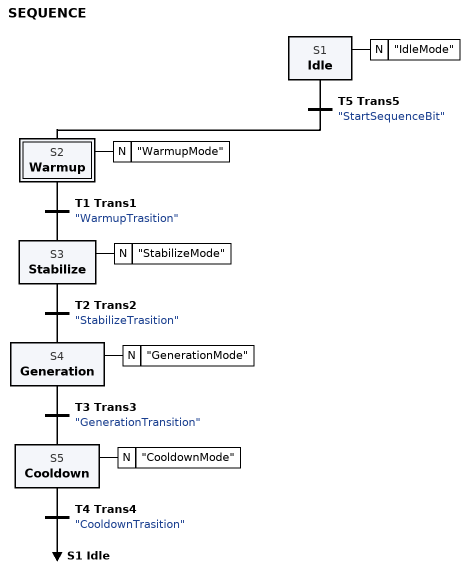
   // sequencer 1
   STEP Idle:   // S1, max time T#10S, warning time T#7S
              N    "IdleMode"
   END_STEP
   TRANSITION Trans5 FROM Idle TO Warmup   // T5
      := "StartSequenceBit";
   END_TRANSITION
   INITIAL_STEP Warmup:   // S2, max time T#10S, warning time T#7S
              N    "WarmupMode"
   END_STEP
   TRANSITION Trans1 FROM Warmup TO Stabilize   // T1
      := "WarmupTrasition";
   END_TRANSITION
   STEP Stabilize:   // S3, max time T#10S, warning time T#7S
              N    "StabilizeMode"
   END_STEP
   TRANSITION Trans2 FROM Stabilize TO Generation   // T2
      := "StabilizeTrasition";
   END_TRANSITION
   STEP Generation:   // S4, max time T#10S, warning time T#7S
              N    "GenerationMode"
   END_STEP
   TRANSITION Trans3 FROM Generation TO Cooldown   // T3
      := "GenerationTransition";
   END_TRANSITION
   STEP Cooldown:   // S5, max time T#10S, warning time T#7S
              N    "CooldownMode"
   END_STEP
   TRANSITION Trans4 FROM Cooldown TO Idle   // T4, jump
      := "CooldownTrasition";
   END_TRANSITION
END_FUNCTION_BLOCK

FUNCTION_BLOCK "HOURMETER_LAD"   // FB19, LAD
{ S7_Optimized_Access := 'TRUE' }
VERSION : 0.1
   VAR
      accum_elapsed : Time;
      OS1 : Bool;
      MinuteTimedDown : Bool;
      HourCountedDown : Bool;
      OS2 : Bool;
      OS3 : Bool;
      DayCountedDown : Bool;
      resettime : Time;
      OS4 : Bool;
      resetrto : Bool;
      minutecounterreset : Bool;
      hourcounterreset : Bool;
   END_VAR
   VAR_TEMP
      resethourmetertrigger : Bool;
   END_VAR
   VAR_TEMP   // added for the SCL form of the ladder/FBD networks
      _w1 : Bool;
      _w2 : Bool;
      _w3 : Bool;
   END_VAR
BEGIN

REGION Network 1
